FUNCTION_BLOCK "LSim_Lagging"   // FB59, SCL
{ S7_Optimized_Access := 'TRUE' }
VERSION : 2.02
   VAR_INPUT
      input : Real;   // input signal
   END_VAR
   VAR_OUTPUT
      output : Real;   // output signal
   END_VAR
   VAR_IN_OUT
      delayCycles : UInt;   // number of cycles the input signal is delayed (if #delayCycles > #MAX then #delayCycles = #MAX)
   END_VAR
   VAR
      statDelayStore : Array[0..#MAX] of Real;
      statIndexRead : Int;
      statIndexWrite : Int;
   END_VAR
   VAR CONSTANT
      MAX : Int := 100;   // maximum size of array #statDelayStore
   END_VAR
BEGIN
   //=============================================================================
   //SIEMENS AG
   //(c)Copyright 2017 All Rights Reserved
   //-----------------------------------------------------------------------------
   //Library:       Library for Controlled System Simulation
   //Tested with:   S7-1500 FW V2.0 / S7-1200 FW V4.2
   //Engineering:   STEP 7 V14 Upd2 (TIA Portal)
   //Restrictions:  Cyclic interrupt
   //Requirements:  memory card needed for S7-1500
   //Functionality: Simulation of an Tt-System (Lagging)
   //
   //  F(p) = EXP(-p * delayCycles * cyclic interrupt time)
   //          
   //  Call the simulation in a cyclic interrupt with
   //  cyclic interrupt time at least = tmLag1/10!
   //-----------------------------------------------------------------------------
   //Change log table:
   //Version  Date       Expert in charge                Changes applied
   //02.00.00 03.02.2016 Siemens Industry Online Support Release (STEP 7 V13 SP1)
   //02.00.01 02.03.2017 Siemens Industry Online Support Optimize program code
   //02.00.02 02.03.2017 Siemens Industry Online Support Release (STEP 7 V14)
   //=============================================================================

   // Check Parameters
   IF #delayCycles > #MAX THEN
     #delayCycles := INT_TO_UINT(#MAX);
   ELSE
     #delayCycles := #delayCycles;
   END_IF;

   IF #statIndexWrite < #delayCycles THEN
     #statDelayStore[#statIndexWrite] := #input;   // write input at delayStore indexWrite
     #statIndexRead := #statIndexWrite + 1;
     #output := #statDelayStore[#statIndexRead];   // read output from delayStore indexWrite + 1
     #statIndexWrite := #statIndexWrite + 1;       // increment delayStore indexWrite
   ELSE // maximum reached
     #statDelayStore[#statIndexWrite] := #input;   // write input at delayStore maximum
     #statIndexRead := 0;                          // set indexRead to beginning
     #output := #statDelayStore[#statIndexRead];   // read output from delayStore indexRead
     #statIndexWrite := 0;                         // set indexWrite to beginning
   END_IF;
END_FUNCTION_BLOCK

FUNCTION_BLOCK "LSim_DT1"   // FB60, SCL
{ S7_Optimized_Access := 'TRUE' }
VERSION : 2.01
   VAR_INPUT
      calcParam : Bool;   // recalculate with new parameters
      input : Real;   // input signal
      tmLag1 : Real := 2.0;   // time constant T1 [sec]
      tmLag2 : Real := 0.5;   // time constant T2 [sec]
      gain : Real := 1.0;   // gain factor
      cycle : Real := 0.1;   // cyclic time [sec]
      maxOut : Real := 100.0;   // max. output limit
      minOut : Real := -100.0;   // min. output limit
      reset : Bool;   // resets all relevant parameters to ‘0’ including the output
   END_VAR
   VAR_OUTPUT
      error : Bool;   // error (#tmLag1 <= 0)
      status : Word;   // status (if #tmLag1 <= 0 then status = 16#8001)
      maxReached : Bool;   // output has reached max. limit
      minReached : Bool;   // output has reached min. limit
      output : Real;   // output signal (if #error = FALSE)
   END_VAR
   VAR
      statRxn1 : Real;   // delayed input signal (n-1)
      statRyn1 : Real;   // delayed output signal (n-1)
      statRb0 : Real;
      statRa1 : Real;
      statOverfirst : Bool;
      statOutput : Real;   // output signal
   END_VAR
BEGIN
   //=============================================================================
   //SIEMENS AG
   //(c)Copyright 2017 All Rights Reserved
   //-----------------------------------------------------------------------------
   //Library:       Library for Controlled System Simulation
   //Tested with:   S7-1500 FW V2.0 / S7-1200 FW V4.2
   //Engineering:   STEP 7 V14 Upd2 (TIA Portal)
   //Restrictions:  Cyclic interrupt
   //Requirements:  memory card needed for S7-1500
   //Functionality: Simulation of a DT1-System
   //
   //         gain * tmLag2 * p
   //  F(p) = ------------------------------
   //            (1 + tmLag1*p)
   //          
   //  Call the simulation in a cyclic interrupt with
   //  cyclic interrupt time at least = tmLag1/10!
   //-----------------------------------------------------------------------------
   //Change log table:
   //Version  Date       Expert in charge                Changes applied
   //02.00.00 03.02.2016 Siemens Industry Online Support Release (STEP 7 V13 SP1)
   //02.00.01 02.03.2017 Siemens Industry Online Support Release (STEP 7 V14)
   //=============================================================================

   // check of the parameter
   IF #tmLag1 <= 0 THEN
     #error := true;
     #status := W#16#8001; // parameter error
     #statRxn1 := 0.0;
     #statRyn1 := 0.0;
     #statOutput := 0;
     #output := 0;
     RETURN;
   ELSE
     #error := FALSE;
     #status := W#16#0000;     // no error
   END_IF;

   // calculates the z-parameter for the difference equatation
   IF #calcParam = True OR NOT #statOverfirst THEN 
     // Calculate the z-parameter for the DT1-System
     #statOverfirst := 1;
     #statRa1 := -EXP(-#cycle/#tmLag1);
     #statRb0 := #gain*(#tmLag2/#tmLag1);
   END_IF;

   // reset Memory
   IF #reset = True THEN
     #statRxn1 := 0.0;
     #statRyn1 := 0.0;
     #statOutput:=0;
     #error := false;
     #status := W#16#0000;
   END_IF;

   // save delayed output-signals
   #statRyn1:= #statOutput;

   //  difference equatation for DT1-system
   #statOutput := #input * #statRb0 - #statRxn1* #statRb0 - #statRyn1*#statRa1;

   // save delayed input-signals
   #statRxn1 := #input;

   // max limit of acutating variable
   IF #statOutput > #maxOut THEN
     #statOutput := #maxOut;
     #maxReached := True;
   ELSE
     #maxReached := False;
   END_IF;

   // min limit of acutating variable
   IF #statOutput < #minOut THEN
     #statOutput := #minOut;
     #minReached := True;
   ELSE
     #minReached := False;
   END_IF;

   #output := #statOutput;
END_FUNCTION_BLOCK

FUNCTION_BLOCK "LSim_AllPass1OrdReal"   // FB61, SCL
{ S7_Optimized_Access := 'TRUE' }
VERSION : 2.01
   VAR_INPUT
      calcParam : Bool;   // recalculate with new parameters
      input : Real;   // input signal
      tmLag1 : Real := 2.0;   // time constant T1 [sec]
      gain : Real := 1.0;   // gain factor
      cycle : Real := 0.1;   // cyclic time [sec]
      maxOut : Real := 100.0;   // max. output limit
      minOut : Real;   // min. output limit
      reset : Bool;   // resets all relevant parameters to ‘0’ including the output
   END_VAR
   VAR_OUTPUT
      error : Bool;   // error (#tmLag1 <= 0)
      status : Word;   // status (if #tmLag1 <= 0 then status = 16#8001)
      maxReached : Bool;   // output has reached max. limit
      minReached : Bool;   // output has reached min. limit
      output : Real;   // output signal (if #error = FALSE)
   END_VAR
   VAR
      statRxn1 : Real;   // delayed input signal (n-1)
      statRyn1 : Real;   // delayed output signal (n-1)
      statRb1 : Real;
      statRa1 : Real;
      statOutput : Real;   // output signal
   END_VAR
BEGIN
   //=============================================================================
   //SIEMENS AG
   //(c)Copyright 2017 All Rights Reserved
   //-----------------------------------------------------------------------------
   //Library:       Library for Controlled System Simulation
   //Tested with:   S7-1500 FW V2.0 / S7-1200 FW V4.2
   //Engineering:   STEP 7 V14 Upd2 (TIA Portal)
   //Restrictions:  Cyclic interrupt
   //Requirements:  memory card needed for S7-1500
   //Functionality: Simulation of an All-Pass 1. Order with real p-Poles
   //
   //         gain * (1 - tmLag1*p)
   //  F(p) = ---------------------
   //            (1 + tmLag1*p)
   //          
   //  Call the simulation in a cyclic interrupt with
   //  cyclic interrupt time at least = tmLag1/10!
   //-----------------------------------------------------------------------------
   //Change log table:
   //Version  Date       Expert in charge                Changes applied
   //02.00.00 03.02.2016 Siemens Industry Online Support Release (STEP 7 V13 SP1)
   //02.00.01 02.03.2017 Siemens Industry Online Support Release (STEP 7 V14)
   //=============================================================================

   // check of the parameter
   IF #tmLag1 <= 0 THEN
     #error := True;
     #status := W#16#8001;     // Parameter Error
     #statRxn1 := 0.0;
     #statRyn1 := 0.0;
     #statOutput := 0;
     #output := 0;
     RETURN;
   ELSE
     #error := FALSE;
     #status := W#16#0000;     // no error
   END_IF;


   // Z-parameters 
   IF #calcParam = True THEN
   // Calculate z-parameters for allpass filter
      #statRa1 := -EXP(-#cycle/#tmLag1);
      #statRb1 := #gain*(2 + #statRa1);

   END_IF;
   // reset Memory
   IF #reset = True THEN
     #statRxn1 := 0.0;
     #statRyn1 := 0.0;
     #statOutput:=0;
     #error := False;
     #status := W#16#0000;
   END_IF;

   // save delayed output signal 
   #statRyn1:= #statOutput;

   // Differencial Equation of all-pass filter 1. order
   #statOutput := #input * (-#gain) +  #statRxn1* #statRb1 - #statRyn1*#statRa1;

   // save delayed input signals
   #statRxn1 := #input;

   // max limit of acutating variable
   IF #statOutput > #maxOut THEN
     #statOutput := #maxOut;
     #maxReached:= True;
   ELSE
     #maxReached := False;
   END_IF;

   // min limit of acutating variable
   IF #statOutput < #minOut THEN
     #statOutput := #minOut;
     #minReached := True;
   ELSE
     #minReached := False;
   END_IF;

   #output := #statOutput;
END_FUNCTION_BLOCK

FUNCTION_BLOCK "LSim_AllPass2OrdReal"   // FB62, SCL
{ S7_Optimized_Access := 'TRUE' }
VERSION : 2.01
   VAR_INPUT
      calcParam : Bool;   // recalculate with new parameters
      input : Real;   // input signal
      tmLag1 : Real := 2.0;   // time constant T1 [sec]
      tmLag2 : Real := 0.2;   // time constant T2 [sec]
      gain : Real := 1.0;   // gain factor
      cycle : Real := 0.1;   // cyclic time [sec]
      maxOut : Real := 100.0;   // max. output limit
      minOut : Real;   // min. output limit
      reset : Bool;   // resets all relevant parameters to ‘0’ including the output
   END_VAR
   VAR_OUTPUT
      error : Bool;   // error (#tmLag1 <= 0 or #tmLag2 <= 0 or #tmLag2 = #tmLag1)
      status : Word;   // status (if #error = TRUE then status = 16#8001)
      maxReached : Bool;   // output has reached max. limit
      minReached : Bool;   // output has reached min. limit
      output : Real;   // output signal (if #error = FALSE)
   END_VAR
   VAR
      statRxn2 : Real;   // delayed input signal (n-2)
      statRxn1 : Real;   // delayed input signal (n-1)
      statRyn2 : Real;   // delayed output signal (n-2)
      statRyn1 : Real;   // delayed output signal (n-1)
      statRb1 : Real;
      statRb2 : Real;
      statRa1 : Real;
      statRa2 : Real;
      statRe1 : Real;
      statRe2 : Real;
      statRk1 : Real;
      statOverfirst : Bool;
      statOutput : Real;   // output signal
   END_VAR
BEGIN
   //=============================================================================
   //SIEMENS AG
   //(c)Copyright 2017 All Rights Reserved
   //-----------------------------------------------------------------------------
   //Library:       Library for Controlled System Simulation
   //Tested with:   S7-1500 FW V2.0 / S7-1200 FW V4.2
   //Engineering:   STEP 7 V14 Upd2 (TIA Portal)
   //Restrictions:  Cyclic interrupt
   //Requirements:  memory card needed for S7-1500
   //Functionality: Simulation of an All-Pass 2. Order with real p-Poles
   //
   //         gain * (1 - tmLag1*p) * (1 - tmLag2*p)
   //  F(p) = --------------------------------------
   //            (1 + tmLag1*p) * (1 + tmLag2*p)
   //          
   //  Call the simulation in a cyclic interrupt with
   //  cyclic interrupt time at least = tmLag1/10!
   //-----------------------------------------------------------------------------
   //Change log table:
   //Version  Date       Expert in charge                Changes applied
   //02.00.00 03.02.2016 Siemens Industry Online Support Release (STEP 7 V13 SP1)
   //02.00.01 02.03.2017 Siemens Industry Online Support Release (STEP 7 V14)
   //=============================================================================

   // check of the parameter
   IF #tmLag1 <= 0 OR #tmLag2 <= 0 OR #tmLag1 = #tmLag2 THEN
     #error := TRUE;
     #status := W#16#8001;     // Parameter Error
     #statRxn1 := 0.0;
     #statRyn1 := 0.0;
     #statRxn2 := 0.0;
     #statRyn2 := 0.0;
     #statOutput := 0;
     #output := 0;
     RETURN;
   ELSE
     #error := FALSE;
     #status := W#16#0000;     // no error
   END_IF;

   // calculates the z-parameter for the difference equatation
   IF #calcParam = True OR NOT #statOverfirst THEN
   // Calculate z-parameters for oscilating PT2-System
   #statOverfirst:=1;
   #statRe1 := -EXP(-#cycle/#tmLag1);
   #statRe2 := -EXP(-#cycle/#tmLag2);
   #statRk1 := (2* (#tmLag2 + #tmLag1))/(#tmLag2 - #tmLag1);
   #statRa1 := #statRe1 + #statRe2;
   #statRa2 := #statRe1*#statRe2;
   #statRb1 := #gain*(#statRa1+ #statRk1*(#statRe2 - #statRe1));
   #statRb2 := #gain*(#statRa2 -#statRk1*(#statRe2 - #statRe1));
   END_IF;

   // reset memory
   IF #reset = True THEN
     #statRxn1 := 0.0;
     #statRyn1 := 0.0;
     #statRxn2 := 0.0;
     #statRyn2 := 0.0;
     #statOutput:=0;
     #error := False;
     #status := W#16#0000;
   END_IF;

   // save delayed output-signals
   #statRyn2:=#statRyn1;
   #statRyn1:= #statOutput;

   // difference equatation for PT2-system
   #statOutput := #input * #gain +  #statRxn1* #statRb1 + #statRxn2*#statRb2 - #statRyn1*#statRa1 - #statRyn2*#statRa2;

   // save delayed input-signals
   #statRxn2 := #statRxn1;
   #statRxn1 := #input;

   // max limit of acutating variable
   IF #statOutput > #maxOut THEN
     #statOutput := #maxOut;
     #maxReached:= True;
   ELSE
     #maxReached := False;
   END_IF;

   // min limit of acutating variable
   IF #statOutput < #minOut THEN
     #statOutput := #minOut;
     #minReached := True;
   ELSE
     #minReached := False;
   END_IF;

   #output := #statOutput;
END_FUNCTION_BLOCK

FUNCTION_BLOCK "LSim_Valve"   // FB63, FBD
{ S7_Optimized_Access := 'TRUE' }
VERSION : 2.01
// //============================================================================
// //SIEMENS AG
// //(c)Copyright 2017 All Rights Reserved
// //-----------------------------------------------------------------------------
// //Library:       Library for Controlled System Simulation
// //Tested with:   S7-1500 FW V2.0 / S7-1200 FW V4.2
// //Engineering:   STEP 7 V14 Upd2 (TIA Portal)
// //Restrictions:  Cyclic interrupt
// //Requirements:  memory card needed for S7-1500
// //Functionality: Simulation of a valve with adjustable transition time
// //-----------------------------------------------------------------------------
// //Change log table:
// //Version    Date             Expert in charge                               Changes applied
// //02.00.00 03.02.2016 Siemens Industry Online Support Release (STEP 7 V13 SP1)
// //02.00.01 02.03.2017 Siemens Industry Online Support Release (STEP 7 V14)
// //============================================================================
   VAR_INPUT
      inputUp : Bool := false;   // control signal “Open valve”
      inputDn : Bool := false;   // control signal “Close valve”
      inputPer : Int;   // Analog manipulated variable
      perOn : Bool;   // selection switch, whether inputUp/inputDn or inputPer is used (inputPer is used for TRUE)
      perMax : Real := 27648.0;   // upper limit of the analog value of the valve position.
      perMin : Real;   // lower limit of the analog value of the valve position
      realMax : Real := 100.0;   // upper limit of the converted floating-point value for the valve position
      realMin : Real;   // lower limit of the converted floating-point value for the valve position
      transitTime : Real := 20.0;   // traversing time of the value between the end positions
      cycle : Real := 0.1;   // cyclic time [sec]
      reset : Bool := false;   // resets all relevant parameters to ‘0’ including the output
   END_VAR
   VAR_OUTPUT
      output : Real := 0.0;   // calculated valve position (within the “realMin” and “realMax” limits)
      outputPer : Int;   // calculated analog valve position (within the “perMin” and “perMax” limits)
      highLimit : Bool := false;   // simulated upper valve end position reached at highLimit = TRUE
      lowLimit : Bool := false;   // simulated lower valve end position reached at lowLimit = TRUE
   END_VAR
   VAR
      statInput : Real;
      statDelta : Real;
      statOut : Real;
      statHigh : Bool;
      statLow : Bool;
   END_VAR
   VAR_TEMP
      tempReal : Real;
      tempStepWidth : Real;
      tempStepWidthNeg : Real;
      tempBool : Bool;
      tempInputNorm : Real;
      tempUpFlag : Bool;
      tempDnFlag : Bool;
      tempInt : Int;
   END_VAR
   VAR_TEMP   // added for the SCL form of the ladder/FBD networks
      _w1 : Bool;
   END_VAR
BEGIN

REGION Network 1: reset
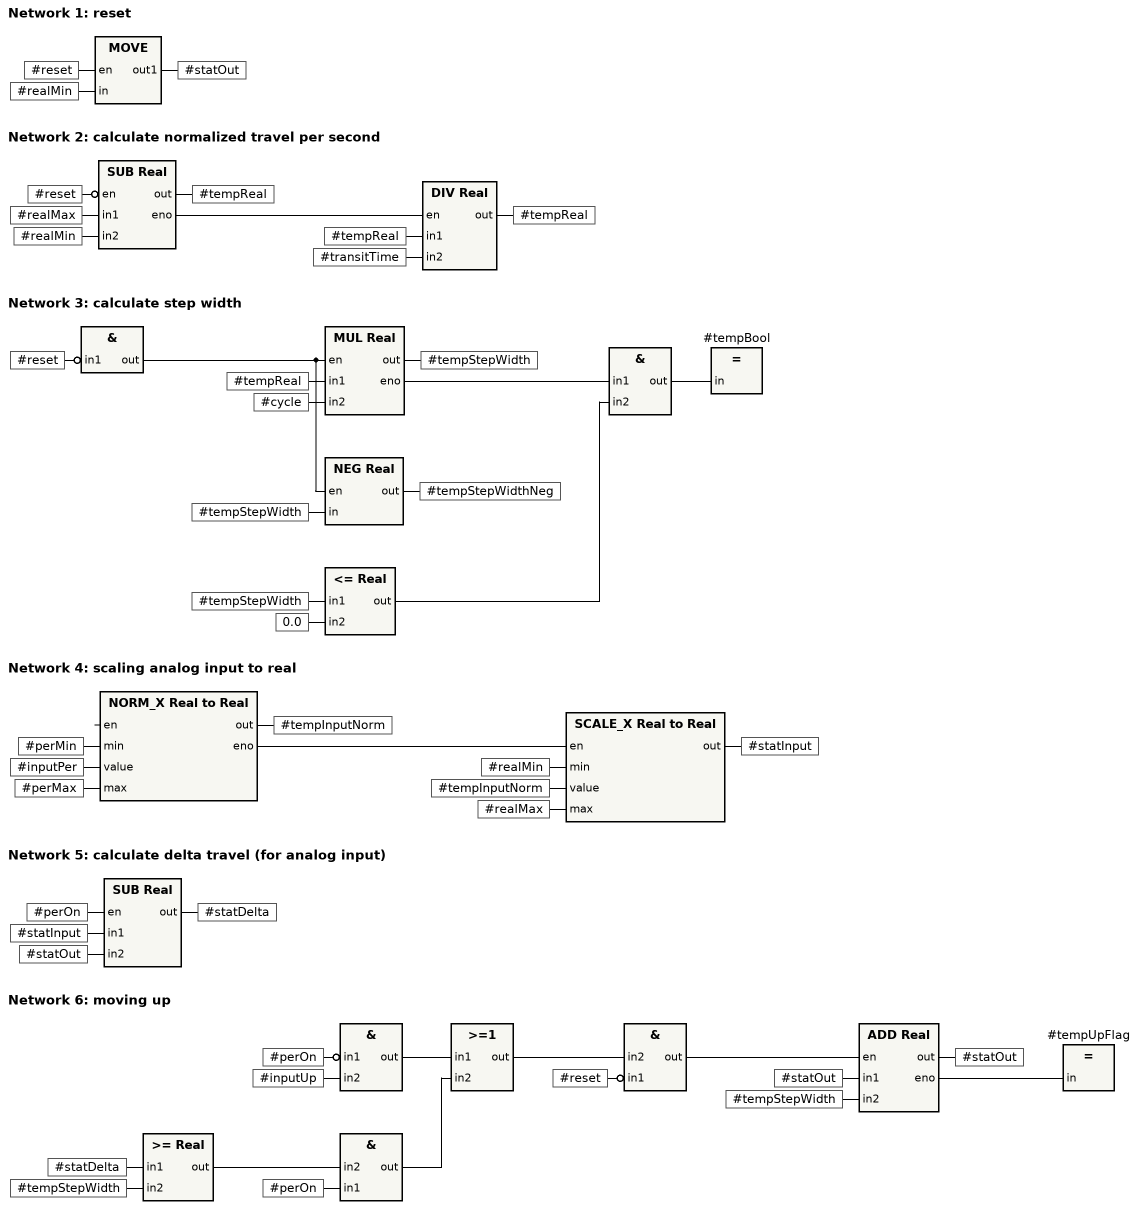
   IF #reset THEN #statOut := #realMin; END_IF;
END_REGION

REGION Network 2: calculate normalized travel per second
   // ENO of a box is taken as its EN; it also drops when the box reports an error
   IF NOT #reset THEN
       #tempReal := #realMax - #realMin;
       #tempReal := #tempReal / #transitTime;
   END_IF;
END_REGION

REGION Network 3: calculate step width
   // ENO of a box is taken as its EN; it also drops when the box reports an error
   IF NOT #reset THEN #tempStepWidth := #tempReal * #cycle; END_IF;
   #tempBool := NOT #reset AND (#tempStepWidth <= 0.0);
   IF NOT #reset THEN #tempStepWidthNeg := -#tempStepWidth; END_IF;
END_REGION

REGION Network 4: scaling analog input to real
   // ENO of a box is taken as its EN; it also drops when the box reports an error
   #tempInputNorm := NORM_X(MIN := #perMin, VALUE := #inputPer, MAX := #perMax);
   #statInput := SCALE_X(MIN := #realMin, VALUE := #tempInputNorm, MAX := #realMax);
END_REGION

REGION Network 5: calculate delta travel (for analog input)
   IF #perOn THEN #statDelta := #statInput - #statOut; END_IF;
END_REGION

REGION Network 6: moving up
   // ENO of a box is taken as its EN; it also drops when the box reports an error
   #_w1 := ((NOT #perOn AND #inputUp) OR ((#statDelta >= #tempStepWidth) AND #perOn)) AND NOT #reset;
   IF #_w1 THEN #statOut := #statOut + #tempStepWidth; END_IF;
   #tempUpFlag := #_w1;
END_REGION

REGION Network 7: checking max. limit
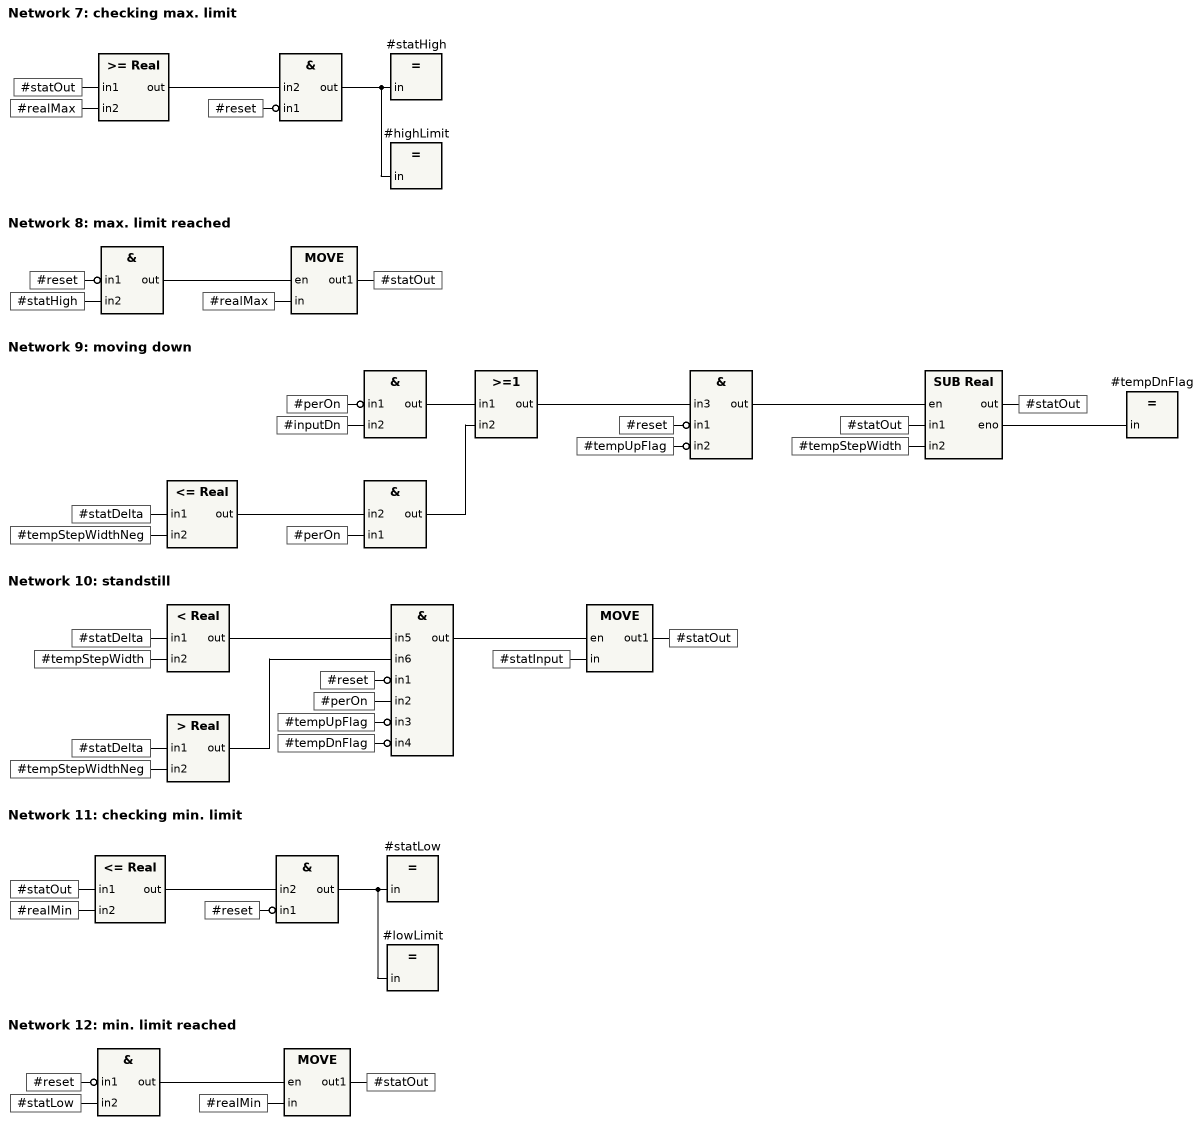
   #statHigh := (#statOut >= #realMax) AND NOT #reset;
   #highLimit := #statHigh;
END_REGION

REGION Network 8: max. limit reached
   IF NOT #reset AND #statHigh THEN #statOut := #realMax; END_IF;
END_REGION

REGION Network 9: moving down
   // ENO of a box is taken as its EN; it also drops when the box reports an error
   #_w1 := ((NOT #perOn AND #inputDn) OR ((#statDelta <= #tempStepWidthNeg) AND #perOn)) AND NOT #reset AND NOT #tempUpFlag;
   IF #_w1 THEN #statOut := #statOut - #tempStepWidth; END_IF;
   #tempDnFlag := #_w1;
END_REGION

REGION Network 10: standstill
   IF (#statDelta < #tempStepWidth) AND (#statDelta > #tempStepWidthNeg) AND NOT #reset AND #perOn AND NOT #tempUpFlag AND NOT #tempDnFlag THEN
       #statOut := #statInput;
   END_IF;
END_REGION

REGION Network 11: checking min. limit
   #statLow := (#statOut <= #realMin) AND NOT #reset;
   #lowLimit := #statLow;
END_REGION

REGION Network 12: min. limit reached
   IF NOT #reset AND #statLow THEN #statOut := #realMin; END_IF;
END_REGION

REGION Network 13: output and scaling to analog
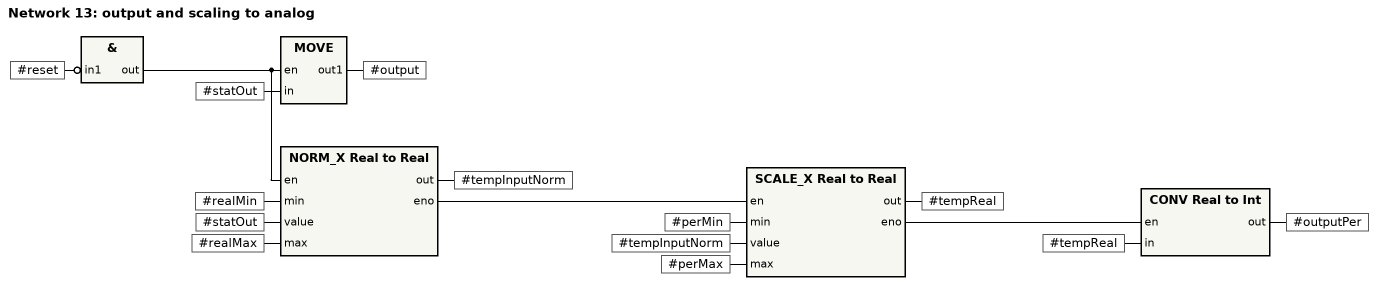
   // ENO of a box is taken as its EN; it also drops when the box reports an error
   IF NOT #reset THEN
       #output := #statOut;
       #tempInputNorm := NORM_X(MIN := #realMin, VALUE := #statOut, MAX := #realMax);
       #tempReal := SCALE_X(MIN := #perMin, VALUE := #tempInputNorm, MAX := #perMax);
       #outputPer := REAL_TO_INT(#tempReal);
   END_IF;
END_REGION
END_FUNCTION_BLOCK

FUNCTION_BLOCK "LSim_PT3HeatCool"   // FB64, SCL
{ S7_Optimized_Access := 'TRUE' }
VERSION : 2.01
   VAR_INPUT
      inputHeat : Real;   // input variable heating
      inputCool : Real;   // input variable cooling
      disturbHeat : Real;   // disturbance variable heating (additional to "inputHeat")
      disturbCool : Real;   // disturbance variable cooling (additional to "inputCool")
      ambTemp : Real := 20.0;   // ambient temperature
      gainHeat : Real := 1.5;   // proportional gain heating
      gainCool : Real := 3.0;   // proportional gain cooling
      tmLag1Heat : Real := 60.0;   // time lag 1 heating [s]
      tmLag2Heat : Real := 10.0;   // time lag 2 heating [s]
      tmLag3Heat : Real;   // time lag 3 heating [s]
      tmLag1Cool : Real := 60.0;   // time lag 1 cooling [s]
      tmLag2Cool : Real := 10.0;   // time lag 2 cooling [s]
      tmLag3Cool : Real;   // time lag 3 cooling [s]
      cycle : Real := 0.1;   // sample time [s]
   END_VAR
   VAR_OUTPUT
      output : Real;   // output variable
   END_VAR
   VAR_IN_OUT
      reset : Bool;   // complete restart
   END_VAR
   VAR
      statFback1 : Array[0..1] of Real;   // feedback value 1 heating/cooling
      statFback2 : Array[0..1] of Real;   // feedback value 2 heating/cooling
      statFback3 : Array[0..1] of Real;   // feedback value 3 heating/cooling
   END_VAR
   VAR_TEMP
      tempHvar : Real;   // helper
      tempCycleR : Real;   // sampling time
      tempTmLag1R : Real;   // delay time 1
      tempTmLag2R : Real;   // delay time 2
      tempTmLag3R : Real;   // delay time 3
      tempIndex : Int;   // control variable
      tempOutvNew : Array[0..1] of Real;   // new output value heating/cooling
   END_VAR
BEGIN
   //=============================================================================
   //SIEMENS AG
   //(c)Copyright 2017 All Rights Reserved
   //-----------------------------------------------------------------------------
   //Library:       Library for Controlled System Simulation
   //Tested with:   S7-1500 FW V2.0 / S7-1200 FW V4.2
   //Engineering:   STEP 7 V14 Upd2 (TIA Portal)
   //Restrictions:  Cyclic interrupt
   //Requirements:  memory card needed for S7-1500
   //Functionality: Simulation of an PT3-system with heating and cooling input
   //-----------------------------------------------------------------------------
   //Change log table:
   //Version  Date       Expert in charge                Changes applied
   //02.00.00 03.02.2016 Siemens Industry Online Support Release (STEP 7 V13 SP1)
   //02.00.01 02.03.2017 Siemens Industry Online Support Release (STEP 7 V14)
   //=============================================================================
   #tempOutvNew[0] := (#inputHeat + #disturbHeat) * #gainHeat;
   #tempOutvNew[1] := (#inputCool + #disturbCool) * #gainCool;

   IF #reset
   THEN
     //restart

     //write output parameters
     #output := #tempOutvNew[0] - #tempOutvNew[1] + #ambTemp;

     //write static local variables
     FOR #tempIndex := 0 TO 1 DO
       #statFback1[#tempIndex] := #tempOutvNew[#tempIndex];
       #statFback2[#tempIndex] := #statFback1[#tempIndex];
       #statFback3[#tempIndex] := #statFback2[#tempIndex];
     END_FOR;

     #reset := FALSE;
   ELSE
     //smoothing  
     #tempCycleR := #cycle;
     IF #tempCycleR < 0.001
     THEN
       //low limit sampling time
       #tempCycleR := 0.001;
     END_IF;

     FOR #tempIndex := 0 TO 1 DO

       IF #tempIndex = 0
       THEN
         #tempTmLag1R := #tmLag1Heat;
         #tempTmLag2R := #tmLag2Heat;
         #tempTmLag3R := #tmLag3Heat;
       ELSE
         #tempTmLag1R := #tmLag1Cool;
         #tempTmLag2R := #tmLag2Cool;
         #tempTmLag3R := #tmLag3Cool;
       END_IF;

       //1.delay
       IF #tempTmLag1R >= #tempCycleR * 0.5
       THEN
         #tempHvar := #tempCycleR / (2.0 * #tempTmLag1R + #tempCycleR);
         #tempHvar := (#tempOutvNew[#tempIndex] - #statFback1[#tempIndex]) * #tempHvar;
         //calculate new output value
         #tempOutvNew[#tempIndex] := #statFback1[#tempIndex] + #tempHvar;
         //calculate new feedback value
         #statFback1[#tempIndex] := #statFback1[#tempIndex] + 2.0 * #tempHvar;
       ELSE  //----------------------------------- implicit PT1
         #tempHvar := #tempCycleR / (#tempTmLag1R + #tempCycleR);
         //calculate new feedback value
         #statFback1[#tempIndex] := #statFback1[#tempIndex] + (#tempOutvNew[#tempIndex] - #statFback1[#tempIndex]) * #tempHvar;
         //calculate new output value
         #tempOutvNew[#tempIndex] := #statFback1[#tempIndex];
       END_IF;

       //2.delay heating
       IF #tempTmLag2R >= #tempCycleR * 0.5
       THEN
         #tempHvar := #tempCycleR / (2.0 * #tempTmLag2R + #tempCycleR);
         #tempHvar := (#tempOutvNew[#tempIndex] - #statFback2[#tempIndex]) * #tempHvar;
         //calculate new output value
         #tempOutvNew[#tempIndex] := #statFback2[#tempIndex] + #tempHvar;
         //calculate new feedback value
         #statFback2[#tempIndex] := #statFback2[#tempIndex] + 2.0 * #tempHvar;
       ELSE
         #statFback2[#tempIndex] := #tempOutvNew[#tempIndex];
       END_IF;

       //3.delay heating
       IF #tempTmLag3R >= #tempCycleR * 0.5
       THEN
         #tempHvar := #tempCycleR / (2.0 * #tempTmLag3R + #tempCycleR);
         #tempHvar := (#tempOutvNew[#tempIndex] - #statFback3[#tempIndex]) * #tempHvar;
         //calculate new output value
         #tempOutvNew[#tempIndex] := #statFback3[#tempIndex] + #tempHvar;
         //calculate new feedback value
         #statFback3[#tempIndex] := #statFback3[#tempIndex] + 2.0 * #tempHvar;
       ELSE
         #statFback3[#tempIndex] := #tempOutvNew[#tempIndex];
       END_IF;

     END_FOR;

     #output := #tempOutvNew[0] - #tempOutvNew[1] + #ambTemp;
   END_IF;
END_FUNCTION_BLOCK

// folder: Mawomat_stare/Klasy_FC

FUNCTION "FC301_Timer" : Void   // FC301, SCL
{ S7_Optimized_Access := 'TRUE' }
VERSION : 0.1
   VAR_INPUT
      iTyp : Int;
      bOnOff : Bool;   // Start zliczania timera
      bRst : Bool;   // Reset
      dCzasZad : DWord;   // Czas zadany timera
      timer_1s : Bool;
   END_VAR
   VAR_OUTPUT
      bOk : Bool;   // Bit oznaczajacy odliczanie timera
   END_VAR
   VAR_IN_OUT
      dCzasAkt : DWord;   // Czas aktualnie zliczony przez timer
   END_VAR
BEGIN
   #bOk := 0;
   IF #iTyp = 1 THEN
       IF (#bOnOff AND (NOT #bRst)) THEN
           IF (#dCzasAkt < #dCzasZad) THEN
               #bOk := 0;
               IF #timer_1s = TRUE THEN
                   #dCzasAkt := #dCzasAkt + 1;
               END_IF;
           ELSE
               #dCzasAkt := #dCzasZad;
               #bOk := 1;
           END_IF;
       ELSE
           #dCzasAkt := 0;
       END_IF;
   END_IF;
END_FUNCTION

FUNCTION "FC321_DIO" : Void   // FC321, SCL
{ S7_Optimized_Access := 'TRUE' }
VERSION : 0.1
   VAR_INPUT
      Nr_Ost_Elementu : Int;   // Numer ostatniego elementu, dla ktorego wykonywana jest klasa
      Nr_Plc : Byte;
   END_VAR
   VAR_TEMP
      i : Int;
   END_VAR
BEGIN
   FOR #i := 1 TO #Nr_Ost_Elementu BY 1 DO
      REGION Opisy bitow sygnalow: bRoz,bSym,bSt,bSt_1,bTrP

                       //bRoz - ROZKAZ OPERATORA - DB321.DBW10 - WORD
                       //bRozB1
                       //"DB321_DIO".DIO[#i].bRoZB1.%X0 - Tryb pracy: 0-Zdalny reczny; 1-Zdalny auto
                       //"DB321_DIO".DIO[#i].bRoZB1.%X1 - Symulacja wejsc urz: 0-Wylaczona; 1-Zalaczona
                       //"DB321_DIO".DIO[#i].bRoZB1.%X2 - Praca z wyjsciami urz: 0-Wylaczona; 1-Zalaczona
                       //"DB321_DIO".DIO[#i].bRoZB1.%X3 - Sterowanie urz. w tr. Zdalnym-Man: 0-Wylacz; 1-Zalacz
                       //"DB321_DIO".DIO[#i].bRoZB1.%X4 - Sterowanie kier. w tr. Zdalnym-Man: 0-Lewa; 1-Prawo
                       //"DB321_DIO".DIO[#i].bRoZB1.%X5-X7 - Rezerwa
                       //bRozB2
                       //"DB321_DIO".DIO[#i].bRoZB2.%X0 - Kasuj awarie (impuls)
                       //"DB321_DIO".DIO[#i].bRoZB2.%X1-X7 - Rezerwa (impuls)
                       //
                       //bSym - SYM WEJSCIA - DB321.DBW12 - WORD
                       //"DB321_DIO".DIO[#i].bSym.%X0 - Aktywacja urz. w systemie (ustawiany tylko z programu)
                       //"DB321_DIO".DIO[#i].bSym.%X1 - Sterowanie urz. w tr. Zdalnym-Auto: 0-Wylacz; 1-Zalacz
                       //"DB321_DIO".DIO[#i].bSym.%X2-X4 - Rezerwa
                       //"DB322_DV1".DV1[#i].bSym.%X5 - Tryb sterowania: 0-Zdalne z PC; 1-Lokalne z elewacji szafy
                       //"DB322_DV1".DV1[#i].bSym.%X6 - Tryb remontowy (z wylacznika): 0-Brak; 1-Aktywny
                       //"DB321_DIO".DIO[#i].bSym.%X7 - Awaria zewnetrzna: 0-Brak; 1-Aktywny
                       //"DB321_DIO".DIO[#i].bSym.%X8 - Blokada zmiany tr. zdalnego z Auto na Man: 0-Brak; 1-Aktywna
                       //"DB321_DIO".DIO[#i].bSym.%X9-X15 - Rezerwa
                       //
                       //bSt_Tryb - STAN - DB321.DBW14 - WORD
                       //"DB321_DIO".DIO[#i].bSt_Tryb.%X0-X1 - Awaria rezerwa
                       //"DB321_DIO".DIO[#i].bSt_Tryb.%X2 - Awaria zewnetzrna: 0-Nieaktywna; 1-Aktywna
                       //"DB321_DIO".DIO[#i].bSt_Tryb.%X3-X7 - Awaria rezerwa
                       //"DB321_DIO".DIO[#i].bSt_Tryb.%X8 - Urzadzenie aktywowane
                       //"DB321_DIO".DIO[#i].bSt_Tryb.%X9 - Blokada zmaiany tr. zdalnego z Auto na Man: 0-Brak; 1-Aktywna
                       //"DB321_DIO".DIO[#i].bSt_Tryb.%X10-X11 - Awaria rezerwa
                       //"DB321_DIO".DIO[#i].bSt_Tryb.%X12 - Symulacja wejsc urzadzenia: 0-Wylaczona; 1-Zalaczona
                       //"DB321_DIO".DIO[#i].bSt_Tryb.%X13 - Praca z wyjsciami urzadzenia: 0-Wylaczona; 1-Zalaczona
                       //"DB321_DIO".DIO[#i].bSt_Tryb.%X14 - Stan urzadzenia: 0-Brak odliczania czasu do otwarcia 1-Odliczanie
                       //"DB321_DIO".DIO[#i].bSt_Tryb.%X15 - Stan urzadzenia: 0-Brak odliczania czasu do zamkniecia 1-Odliczanie
                       //
                       //bSt_Urz - STAN - DB321.DBW16 - INT
                       //"DB321_DIO".DIO[#i].bSt_Urz.%X0 - STAN(1)- Awaria zbiorcza 1-Aktywna; 0-Brak aktywnosci obiektu
                       //"DB321_DIO".DIO[#i].bSt_Urz.%X1 - STAN(2)- Urzadzenie: 1-Zamkniete; 0-Inny stan
                       //"DB321_DIO".DIO[#i].bSt_Urz.%X2 - STAN(4)- Urzadzenie: 1-Otwieraniee; 0-Inny stan
                       //"DB321_DIO".DIO[#i].bSt_Urz.%X3 - STAN(8)- Urzadzenie: 1-Otwarte; 0-Inny stan
                       //"DB321_DIO".DIO[#i].bSt_Urz.%X4 - STAN(16)- Urzadzenie: 1-Zamykanie; 0-Inny stan
                       //"DB321_DIO".DIO[#i].bSt_Urz.%X5 - STAN(32)- Urzadzenie: 1-Odliczanie czasu zwloki awarii; 0-Inny stan
                       //"DB321_DIO".DIO[#i].bSt_Urz.%X6-X7 - STAN- Stan rezerwa
                       //
                       //bTrP - TRYB PRACY - DB321.DBW17 - INT
                       //"DB321_DIO".DIO[#i].bTrP.%X0 - TRYB PRACY(1) - Tryb Remontowy(1): 1-Rezerwa; 0-Brak aktywnosci obiektu
                       //"DB321_DIO".DIO[#i].bTrP.%X1 - Tryb PRACY(2): Rezerwa
                       //"DB321_DIO".DIO[#i].bTrP.%X2 - TRYB PRACY(4) - Tryb Sterowania Zdalnego: 1-Zdalny Reczny; 0-Inny stan
                       //"DB321_DIO".DIO[#i].bTrP.%X3 - TRYB PRACY(8) - Tryb Sterowania Zdalnego: 1-Zdalny Automatyczny; 0-Inny stan
                       //"DB321_DIO".DIO[#i].bTrP.%X4-X7 - Tryb PRACY(16)(32)(64)(128): Rezerwa
                   END_REGION
      REGION Przepisanie danych do obiektu
                       "DB321_DIO".DIO[#i].yNrID := #i;
                       "DB321_DIO".DIO[#i].yNrPLC := #Nr_Plc;
                   END_REGION
           REGION Warunek na wykonanie funkcji
          "DB321_DIO".DIO[#i].bSym.%X0 := "DB321_DIO".DIO[#i].bWeAkt;
          IF "DB321_DIO".DIO[#i].bWeAkt = 0 THEN //Akcja przy deaktywowaniu obiektu
                  "DB321_DIO".DIO[#i].bWeZalAuto := 0;
                  "DB321_DIO".DIO[#i].bWeAwrZ := 0;
                  "DB321_DIO".DIO[#i].bWeBlZmAuto := 0;
                  "DB321_DIO".DIO[#i].bRoZB1 := 0;
                  "DB321_DIO".DIO[#i].bRoZB2 := 0;
                  "DB321_DIO".DIO[#i].bSym := 0;
                  "DB321_DIO".DIO[#i].bSt_Tryb := 0;
                  "DB321_DIO".DIO[#i].bSt_Urz := 0;
                  "DB321_DIO".DIO[#i].bTrP := 0;
                  "DB321_DIO".DIO[#i].bWySter := 0;
                  "DB321_DIO".DIO[#i].bWyRst := 0;
                  "DB321_DIO".DIO[#i].bWeTrRem := 0;
                  "DB321_DIO".DIO[#i].bWeTrLok := 0;
              ELSE
                   REGION Program funckji
                       REGION Symulacja wejsc - przepisywanie wartosci wejsciowych, gdy nie ma symulacji oprocz bWeAkt
                           IF "DB321_DIO".DIO[#i].bSt_Tryb.%X12 = 0 THEN
                               "DB321_DIO".DIO[#i].bSym.%X1 := "DB321_DIO".DIO[#i].bWeZalAuto;
                               "DB321_DIO".DIO[#i].bSym.%X7 := "DB321_DIO".DIO[#i].bWeAwrZ;
                               "DB321_DIO".DIO[#i].bSym.%X8 := "DB321_DIO".DIO[#i].bWeBlZmAuto;
                               "DB321_DIO".DIO[#i].bSym.%X5 := "DB321_DIO".DIO[#i].bWeTrLok;
                               "DB321_DIO".DIO[#i].bSym.%X6 := "DB321_DIO".DIO[#i].bWeTrRem;
                           END_IF;
                       END_REGION
                       REGION Okreslenie stanow
                           "DB321_DIO".DIO[#i].bSt_Tryb.%X8 := "DB321_DIO".DIO[#i].bWeAkt;
                           "DB321_DIO".DIO[#i].bSt_Tryb.%X9 := (("DB321_DIO".DIO[#i].bSym.%X8 AND "DB321_DIO".DIO[#i].bSt_Tryb.%X12) OR ("DB321_DIO".DIO[#i].bWeBlZmAuto AND NOT "DB321_DIO".DIO[#i].bSt_Tryb.%X12));
                           "DB321_DIO".DIO[#i].bSt_Tryb.%X12 := "DB321_DIO".DIO[#i].bRoZB1.%X1;
                           "DB321_DIO".DIO[#i].bSt_Tryb.%X13 := "DB321_DIO".DIO[#i].bRoZB1.%X2;
                       END_REGION
                       REGION Filtracja
                           REGION Timer 1 - opoznienie zalaczenia
                               "DB321_DIO".DIO[#i].bTmr_On_Start := ("DB321_DIO".DIO[#i].bSym.%X1 AND "DB321_DIO".DIO[#i].bSt_Tryb.%X12) OR ("DB321_DIO".DIO[#i].bWeZalAuto AND NOT "DB321_DIO".DIO[#i].bSt_Tryb.%X12);
                               "DB321_DIO".DIO[#i].bTmr_Off_Start := NOT (("DB321_DIO".DIO[#i].bSym.%X1 AND "DB321_DIO".DIO[#i].bSt_Tryb.%X12) OR ("DB321_DIO".DIO[#i].bWeZalAuto AND NOT "DB321_DIO".DIO[#i].bSt_Tryb.%X12));
                               "FC301_Timer"(iTyp := 1,
                                             bOnOff := "DB321_DIO".DIO[#i].bTmr_On_Start,
                                             bRst := 0,
                                             dCzasZad := "DB321_DIO".DIO[#i].yCzZadOpzZal,
                                             timer_1s := "imp1s",
                                             bOk => "DB321_DIO".DIO[#i].bTmr_On_Ok,
                                             dCzasAkt := "DB321_DIO".DIO[#i].yCzAktOpzZal);
                               "FC301_Timer"(iTyp := 1,
                                             bOnOff := "DB321_DIO".DIO[#i].bTmr_Off_Start,
                                             bRst := 0,
                                             dCzasZad := "DB321_DIO".DIO[#i].yCzZadOpzWyl,
                                             timer_1s := "imp1s",
                                             bOk => "DB321_DIO".DIO[#i].bTmr_Off_Ok,
                                             dCzasAkt := "DB321_DIO".DIO[#i].yCzAktOpzWyl);

                           END_REGION
                           REGION Efekt dzialania timerow
                               IF "DB321_DIO".DIO[#i].bTmr_On_Ok THEN
                                   "DB321_DIO".DIO[#i].bHlp187 := 1;
                               END_IF;
                               IF "DB321_DIO".DIO[#i].bTmr_Off_Ok OR "DB321_DIO".DIO[#i].bSt_Urz = 1 THEN
                                   "DB321_DIO".DIO[#i].bHlp187 := 0;
                               END_IF;
                           END_REGION
                           REGION Stany zaworu przy odliczaniu czasu
                               "DB321_DIO".DIO[#i].bSt_Tryb.%X14 := "DB321_DIO".DIO[#i].bTmr_On_Start AND NOT "DB321_DIO".DIO[#i].bTmr_On_Ok;

                               "DB321_DIO".DIO[#i].bSt_Tryb.%X15 := ("DB321_DIO".DIO[#i].bTmr_Off_Start AND NOT "DB321_DIO".DIO[#i].bTmr_Off_Ok);

                           END_REGION


                       END_REGION
                       REGION Generowanie sygnalu alarmu - Brak generowania sygnalu alarmu od potwierdzen
                           //Ustawianie i kasowanie sygnalu awarii
                           IF ("DB321_DIO".DIO[#i].bWeAwrZ AND NOT "DB321_DIO".DIO[#i].bSt_Tryb.%X12) OR ("DB321_DIO".DIO[#i].bSym.%X7 AND  "DB321_DIO".DIO[#i].bSt_Tryb.%X12) THEN
                               "DB321_DIO".DIO[#i].bSt_Tryb.%X2 := 1;
                           END_IF;
                           IF "DB321_DIO".DIO[#i].bRoZB2.%X0 THEN
                               "DB321_DIO".DIO[#i].bSt_Tryb := 0
                               ;
                           END_IF;


                       END_REGION
                       REGION Tryb pracy i sterowanie wyjsciem
                           REGION Przepisanie potwierdzen na sterowanie reczny gdy tryb zdalny-auto
                               // Przypadek gdy ktos z wlaczonym automatycznie urz. przechodzi na tryb zdalny-reczn
                               IF "DB321_DIO".DIO[#i].bTrP.%X3 THEN
                                   "DB321_DIO".DIO[#i].bRoZB1.%X3 := (("DB321_DIO".DIO[#i].bWeZalAuto AND NOT "DB321_DIO".DIO[#i].bSt_Tryb.%X12) OR ("DB321_DIO".DIO[#i].bSym.%X1 AND "DB321_DIO".DIO[#i].bSt_Tryb.%X12));
                               END_IF; 
                               IF "DB321_DIO".DIO[#i].bTrP.%X3 AND "DB321_DIO".DIO[#i].bSt_Tryb.%X9 THEN
                                   "DB321_DIO".DIO[#i].bRoZB1.%X0 := 1
                                   ;
                               END_IF;
                           END_REGION
                           REGION Okreslenie trybu pracy wyjscia
                               IF "DB321_DIO".DIO[#i].bRoZB1.%X0 AND NOT "DB321_DIO".DIO[#i].bSt_Tryb.%X9 THEN
                                   "DB321_DIO".DIO[#i].bTrP := 8
                                   ;
                               END_IF;
                               IF NOT "DB321_DIO".DIO[#i].bRoZB1.%X0 THEN
                                   "DB321_DIO".DIO[#i].bTrP := 4
                                   ;
                               END_IF;
                               IF ("DB321_DIO".DIO[#i].bWeTrLok AND NOT "DB321_DIO".DIO[#i].bSt_Tryb.%X12) OR ("DB321_DIO".DIO[#i].bSym.%X5 AND "DB321_DIO".DIO[#i].bSt_Tryb.%X12) THEN
                                   "DB321_DIO".DIO[#i].bTrP := 2
                                   ;
                               END_IF;

                               IF ("DB321_DIO".DIO[#i].bWeTrRem AND NOT "DB321_DIO".DIO[#i].bSt_Tryb.%X12) OR ("DB321_DIO".DIO[#i].bSym.%X6 AND "DB321_DIO".DIO[#i].bSt_Tryb.%X12) THEN
                                   "DB321_DIO".DIO[#i].bTrP := 1
                                   ;
                               END_IF;
                           END_REGION
                           REGION Sterowanie wyjsciem
                               IF NOT "DB321_DIO".DIO[#i].bLatch THEN
                                   "DB321_DIO".DIO[#i].bHlp186 := "DB321_DIO".DIO[#i].bSt_Urz <> 1 AND (("DB321_DIO".DIO[#i].bTrP.%X3 AND "DB321_DIO".DIO[#i].bHlp187) OR ("DB321_DIO".DIO[#i].bTrP.%X2 AND "DB321_DIO".DIO[#i].bRoZB1.%X3));
                               ELSIF "DB321_DIO".DIO[#i].bRoZB2.%X0 THEN
                                   "DB321_DIO".DIO[#i].bHlp186 := 0;
                               ELSIF "DB321_DIO".DIO[#i].bLatch AND "DB321_DIO".DIO[#i].bSt_Urz <> 1 AND (("DB321_DIO".DIO[#i].bTrP.%X3 AND "DB321_DIO".DIO[#i].bHlp187) OR ("DB321_DIO".DIO[#i].bTrP.%X2 AND "DB321_DIO".DIO[#i].bRoZB1.%X3)) THEN
                                   "DB321_DIO".DIO[#i].bHlp186 := 1;
                               END_IF;

                               "DB321_DIO".DIO[#i].bWySter := "DB321_DIO".DIO[#i].bHlp186 AND "DB321_DIO".DIO[#i].bSt_Tryb.%X13;

                           END_REGION
                           REGION Sterowanie resetem

                               "DB321_DIO".DIO[#i].bWyRst := "DB321_DIO".DIO[#i].bRoZB2.%X0;
                           END_REGION
                           REGION Stan urzadzenia
                               "DB321_DIO".DIO[#i].bSt_Urz := 0;

                               IF "DB321_DIO".DIO[#i].bSt_Tryb.%X2 THEN
                                   "DB321_DIO".DIO[#i].bSt_Urz := 1;  //awaria zbiorcza aktywna
                               ELSE
                                   IF "DB321_DIO".DIO[#i].bHlp186 = 0 THEN
                                       "DB321_DIO".DIO[#i].bSt_Urz := 2; //urzadzenie zamkniete
                                   ELSIF "DB321_DIO".DIO[#i].bHlp186 = 1 THEN
                                       "DB321_DIO".DIO[#i].bSt_Urz := 8; //urzadzenie otwarte
                                   END_IF;
                               END_IF;




                           END_REGION






                       END_REGION
                       REGION Ustawienia koncowe
                           // Samokasowanie sygnalow
                           "DB321_DIO".DIO[#i].bRoZB2 := 0;
                           IF "DB321_DIO".DIO[#i].bAoff = 1 THEN
                               "DB321_DIO".DIO[#i].bWeZalAuto := 0;
                           END_IF;
                       END_REGION
                   END_REGION
               END_IF;
          END_REGION
     END_FOR;
END_FUNCTION

FUNCTION "FC322_DV1" : Void   // FC322, SCL
{ S7_Optimized_Access := 'TRUE' }